(* Logix 5000 project; controller NWGG 1756-L72 rev 35.12; software revision 35.00; part 4 of 19 *)
(* tags used below, declared in another part *)
   DIST_MOVE : ALIAS FOR I3.10;
   DIST_TO_CL : ALIAS FOR I7.2;
   DS_CLEAN_B : ALIAS FOR O13.5;
   DS_DLY_OFF : ALIAS FOR T4[33];
   DS_M : ALIAS FOR O24[1].0;
   DS_M_B : ALIAS FOR B3[101].0;
   DS_MOV_CCW : ALIAS FOR B3[100].13;
   DS_MOV_CW : ALIAS FOR B3[100].12;
   DS_MOVE_SE : ALIAS FOR T4[32];
   DS_POS8 : ALIAS FOR O13.7;
   DS_POS9 : ALIAS FOR O13.8;
   DS_POS_1 : ALIAS FOR I24[0].2;
   DS_POS_10 : ALIAS FOR I24[0].11;
   DS_POS_2 : ALIAS FOR I24[0].3;
   DS_POS_3 : ALIAS FOR I24[0].4;
   DS_POS_4 : ALIAS FOR I24[0].5;
   DS_POS_5 : ALIAS FOR I24[0].6;
   DS_POS_6 : ALIAS FOR I24[0].7;
   DS_POS_7 : ALIAS FOR I24[0].8;
   DS_POS_8 : ALIAS FOR I24[0].9;
   DS_POS_9 : ALIAS FOR I24[0].10;
   DS_SEEK_1 : ALIAS FOR B3[102].1;
   DS_SEEK_10 : ALIAS FOR B3[102].10;
   DS_SEEK_2 : ALIAS FOR B3[102].2;
   DS_SEEK_3 : ALIAS FOR B3[102].3;
   DS_SEEK_4 : ALIAS FOR B3[102].4;
   DS_SEEK_5 : ALIAS FOR B3[102].5;
   DS_SEEK_6 : ALIAS FOR B3[102].6;
   DS_SEEK_7 : ALIAS FOR B3[102].7;
   DS_SEEK_8 : ALIAS FOR B3[102].8;
   DS_SEEK_9 : ALIAS FOR B3[102].9;
   DS_SET_IN : ALIAS FOR N10[0];
   DS_SPOUT_C : ALIAS FOR O24[1].3;
   DS_SPOUT_C1 : ALIAS FOR O24[1].4;
   DS_SPOUT_D : ALIAS FOR I24[0].1;
   DS_SPOUT_D1 : ALIAS FOR O24[1].1;
   DS_SPOUT_D3 : ALIAS FOR B3[101].1;
   DS_SPOUT_U : ALIAS FOR I24[0].0;
   DS_SPOUT_U1 : ALIAS FOR O24[1].2;
   DS_SPOUT_U2 : ALIAS FOR B3[101].2;
   DS_START_M : ALIAS FOR B3[102].11;
   DS_STOP_MO : ALIAS FOR B3[102].0;
   DS_T21 : ALIAS FOR O13.0;
   DS_T22 : ALIAS FOR O13.1;
   DS_T23 : ALIAS FOR O13.9;
   DS_T231 : ALIAS FOR O13.2;
   DS_T24 : ALIAS FOR O13.3;
   DS_T25 : ALIAS FOR O13.4;
   DS_T26 : ALIAS FOR O13.6;
   I24_004_Bit03 : ALIAS FOR I24[4].3;
   I24_004_Bit04 : ALIAS FOR I24[4].4;
   I24_004_Bit05 : ALIAS FOR I24[4].5;
   I24_004_Bit06 : ALIAS FOR I24[4].6;
   I24_004_Bit07 : ALIAS FOR I24[4].7;
   I24_004_Bit08 : ALIAS FOR I24[4].8;
   I24_004_Bit09 : ALIAS FOR I24[4].9;
   I24_004_Bit10 : ALIAS FOR I24[4].10;
   I24_004_Bit11 : ALIAS FOR I24[4].11;
   I24_004_Bit12 : ALIAS FOR I24[4].12;
   I2_000_Bit07 : ALIAS FOR I2.7;
   I2_000_Bit10 : ALIAS FOR I2.10;
   I2_000_Bit13 : ALIAS FOR I2.13;
   I3_000_Bit01 : ALIAS FOR I3.1;
   I3_000_Bit04 : ALIAS FOR I3.4;
   I3_000_Bit07 : ALIAS FOR I3.7;
   O24_005_Bit03 : ALIAS FOR O24[5].3;
   O24_005_Bit04 : ALIAS FOR O24[5].4;
   O24_005_Bit05 : ALIAS FOR O24[5].5;
   O24_005_Bit06 : ALIAS FOR O24[5].6;
   O24_005_Bit07 : ALIAS FOR O24[5].7;
   O24_005_Bit08 : ALIAS FOR O24[5].8;
   O24_005_Bit09 : ALIAS FOR O24[5].9;
   O24_005_Bit10 : ALIAS FOR O24[5].10;
   O24_005_Bit11 : ALIAS FOR O24[5].11;
   O24_005_Bit12 : ALIAS FOR O24[5].12;
   P10_AUTO_S : ALIAS FOR B3[5].10;
   P10_RUN_AU1 : ALIAS FOR B3[4].10;
   P10_SEC_SE : ALIAS FOR B17[1].10;
   P4_RUN_AUT1 : ALIAS FOR B3[4].4;
   P4_SEC_SEL : ALIAS FOR B17[1].4;
   P5_AUTO_SE : ALIAS FOR B3[5].5;
   P5_RUN_AUT1 : ALIAS FOR B3[4].5;
   P5_SEC_SEL : ALIAS FOR B17[1].5;
   P6_AUTO_SE : ALIAS FOR B3[5].6;
   P6_RUN_AUT1 : ALIAS FOR B3[4].6;
   P6_SEC_SEL : ALIAS FOR B17[1].6;
   P7_AUTO_SE : ALIAS FOR B3[5].7;
   P7_RUN_AUT1 : ALIAS FOR B3[4].7;
   P7_SEC_SEL : ALIAS FOR B17[1].7;
   P8_AUTO_SE : ALIAS FOR B3[5].8;
   P8_RUN_AUT1 : ALIAS FOR B3[4].8;
   P8_SEC_SEL : ALIAS FOR B17[1].8;
   P_RESET_AU : ALIAS FOR B3[4].0;
   SYMBOL_ANA : ALIAS FOR N10[1];
   T11_TREAT : ALIAS FOR B3[11].0;
   T12_TREAT : ALIAS FOR B3[12].0;
   T13_TREAT : ALIAS FOR B3[13].0;
   T13C_TREAT : ALIAS FOR B21[70].10;
   T14_TREAT : ALIAS FOR B3[14].0;
   T15_TREAT : ALIAS FOR B3[15].0;
   T16_TREAT : ALIAS FOR B3[16].0;
   T17_TREAT : ALIAS FOR B3[17].0;
   T19C_TREAT : ALIAS FOR B21[71].10;
   T21_TREAT : ALIAS FOR B3[21].0;
   T22_TREAT : ALIAS FOR B3[22].0;
   T23_TREAT : ALIAS FOR B3[23].0;
   T24_TREAT : ALIAS FOR B3[24].0;
   T25_TREAT : ALIAS FOR B3[25].0;
   T26_TREAT : ALIAS FOR B3[26].0;
   T27_TREAT : ALIAS FOR B3[27].0;
   T28_TREAT : ALIAS FOR B3[28].0;
   T29_TREAT : ALIAS FOR B3[29].0;
(* _2_MAIN, continued *)

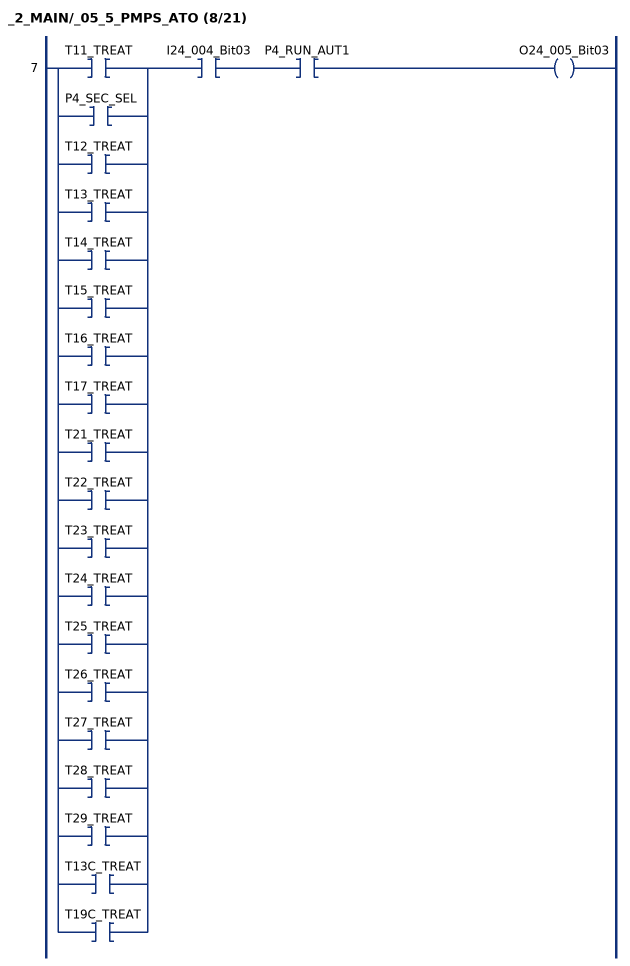
   [picture p56: _2_MAIN/_05_5_PMPS_ATO rungs 7-7]
   7: [XIC(T11_TREAT) ,XIC(P4_SEC_SEL) ,XIC(T12_TREAT) ,XIC(T13_TREAT) ,XIC(T14_TREAT) ,XIC(T15_TREAT) ,XIC(T16_TREAT) ,XIC(T17_TREAT) ,XIC(T21_TREAT) ,XIC(T22_TREAT) ,XIC(T23_TREAT) ,XIC(T24_TREAT) ,XIC(T25_TREAT) ,XIC(T26_TREAT) ,XIC(T27_TREAT) ,XIC(T28_TREAT) ,XIC(T29_TREAT) ,XIC(T13C_TREAT) ,XIC(T19C_TREAT) ]XIC(I24_004_Bit03)XIC(P4_RUN_AUT1)OTE(O24_005_Bit03);
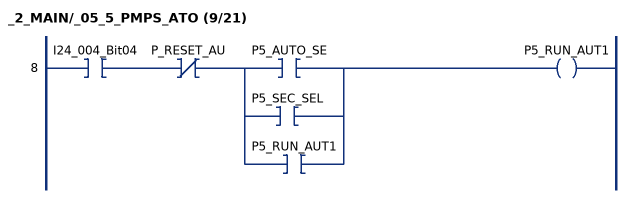
   8: XIC(I24_004_Bit04)XIO(P_RESET_AU)[XIC(P5_AUTO_SE) ,XIC(P5_SEC_SEL) ,XIC(P5_RUN_AUT1) ]OTE(P5_RUN_AUT1);
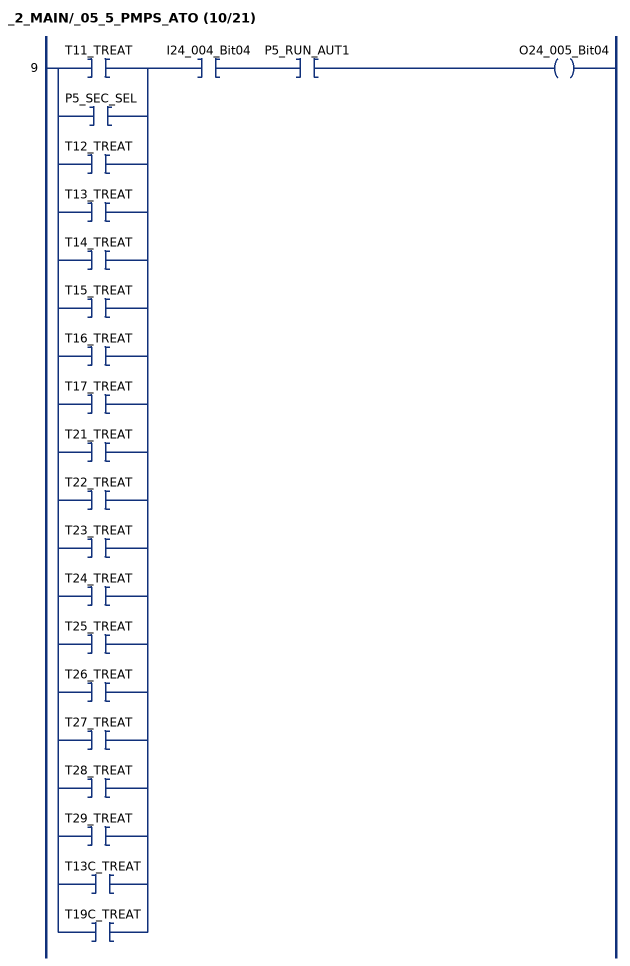
   9: [XIC(T11_TREAT) ,XIC(P5_SEC_SEL) ,XIC(T12_TREAT) ,XIC(T13_TREAT) ,XIC(T14_TREAT) ,XIC(T15_TREAT) ,XIC(T16_TREAT) ,XIC(T17_TREAT) ,XIC(T21_TREAT) ,XIC(T22_TREAT) ,XIC(T23_TREAT) ,XIC(T24_TREAT) ,XIC(T25_TREAT) ,XIC(T26_TREAT) ,XIC(T27_TREAT) ,XIC(T28_TREAT) ,XIC(T29_TREAT) ,XIC(T13C_TREAT) ,XIC(T19C_TREAT) ]XIC(I24_004_Bit04)XIC(P5_RUN_AUT1)OTE(O24_005_Bit04);
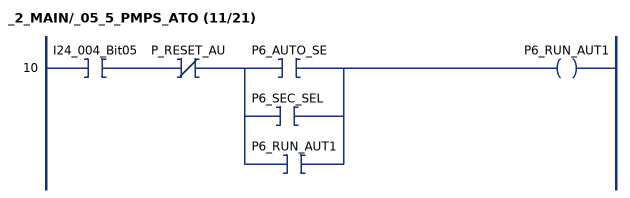
   10: XIC(I24_004_Bit05)XIO(P_RESET_AU)[XIC(P6_AUTO_SE) ,XIC(P6_SEC_SEL) ,XIC(P6_RUN_AUT1) ]OTE(P6_RUN_AUT1);
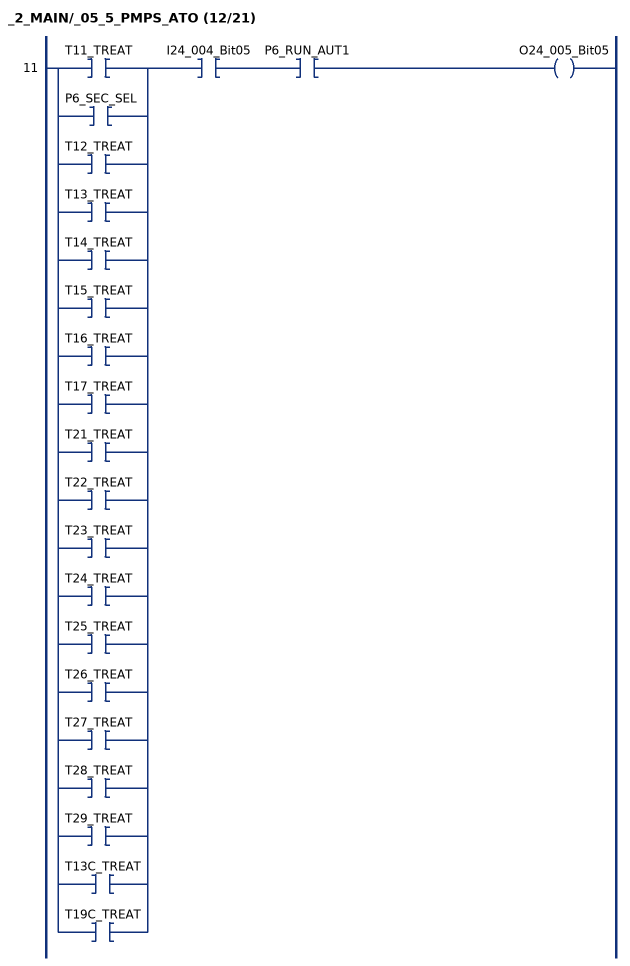
   11: [XIC(T11_TREAT) ,XIC(P6_SEC_SEL) ,XIC(T12_TREAT) ,XIC(T13_TREAT) ,XIC(T14_TREAT) ,XIC(T15_TREAT) ,XIC(T16_TREAT) ,XIC(T17_TREAT) ,XIC(T21_TREAT) ,XIC(T22_TREAT) ,XIC(T23_TREAT) ,XIC(T24_TREAT) ,XIC(T25_TREAT) ,XIC(T26_TREAT) ,XIC(T27_TREAT) ,XIC(T28_TREAT) ,XIC(T29_TREAT) ,XIC(T13C_TREAT) ,XIC(T19C_TREAT) ]XIC(I24_004_Bit05)XIC(P6_RUN_AUT1)OTE(O24_005_Bit05);
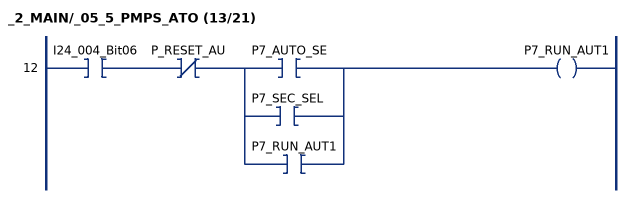
   12: XIC(I24_004_Bit06)XIO(P_RESET_AU)[XIC(P7_AUTO_SE) ,XIC(P7_SEC_SEL) ,XIC(P7_RUN_AUT1) ]OTE(P7_RUN_AUT1);
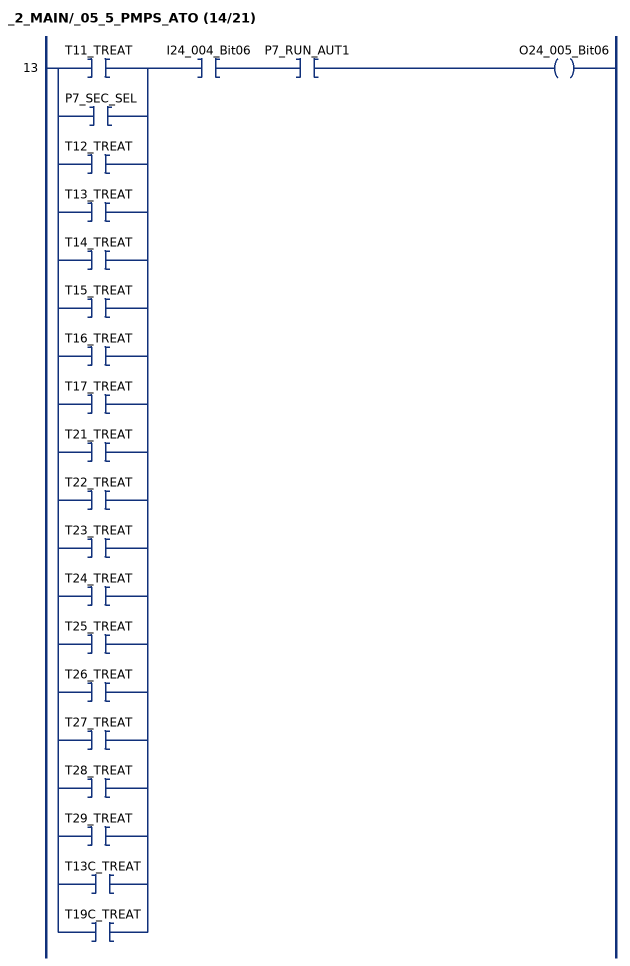
   13: [XIC(T11_TREAT) ,XIC(P7_SEC_SEL) ,XIC(T12_TREAT) ,XIC(T13_TREAT) ,XIC(T14_TREAT) ,XIC(T15_TREAT) ,XIC(T16_TREAT) ,XIC(T17_TREAT) ,XIC(T21_TREAT) ,XIC(T22_TREAT) ,XIC(T23_TREAT) ,XIC(T24_TREAT) ,XIC(T25_TREAT) ,XIC(T26_TREAT) ,XIC(T27_TREAT) ,XIC(T28_TREAT) ,XIC(T29_TREAT) ,XIC(T13C_TREAT) ,XIC(T19C_TREAT) ]XIC(I24_004_Bit06)XIC(P7_RUN_AUT1)OTE(O24_005_Bit06);
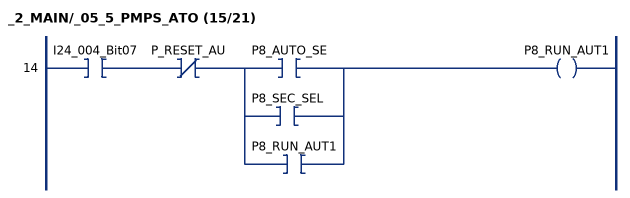
   14: XIC(I24_004_Bit07)XIO(P_RESET_AU)[XIC(P8_AUTO_SE) ,XIC(P8_SEC_SEL) ,XIC(P8_RUN_AUT1) ]OTE(P8_RUN_AUT1);
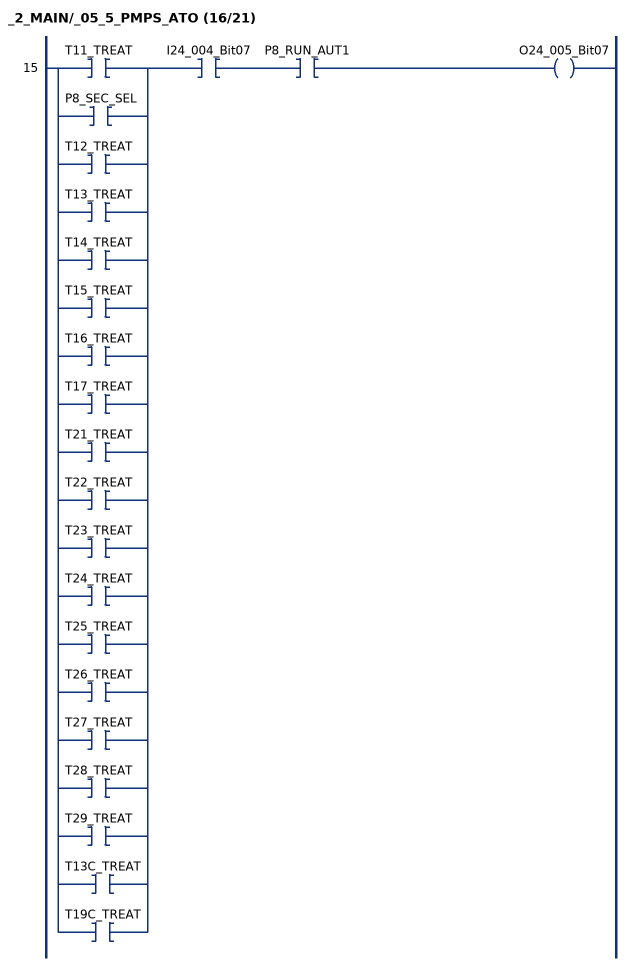
   15: [XIC(T11_TREAT) ,XIC(P8_SEC_SEL) ,XIC(T12_TREAT) ,XIC(T13_TREAT) ,XIC(T14_TREAT) ,XIC(T15_TREAT) ,XIC(T16_TREAT) ,XIC(T17_TREAT) ,XIC(T21_TREAT) ,XIC(T22_TREAT) ,XIC(T23_TREAT) ,XIC(T24_TREAT) ,XIC(T25_TREAT) ,XIC(T26_TREAT) ,XIC(T27_TREAT) ,XIC(T28_TREAT) ,XIC(T29_TREAT) ,XIC(T13C_TREAT) ,XIC(T19C_TREAT) ]XIC(I24_004_Bit07)XIC(P8_RUN_AUT1)OTE(O24_005_Bit07);
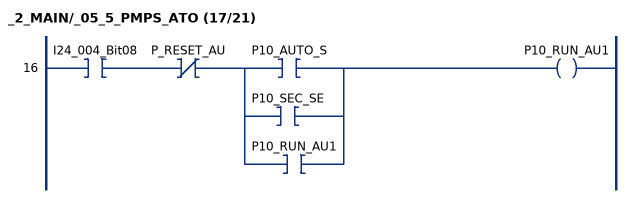
   16: XIC(I24_004_Bit08)XIO(P_RESET_AU)[XIC(P10_AUTO_S) ,XIC(P10_SEC_SE) ,XIC(P10_RUN_AU1) ]OTE(P10_RUN_AU1);
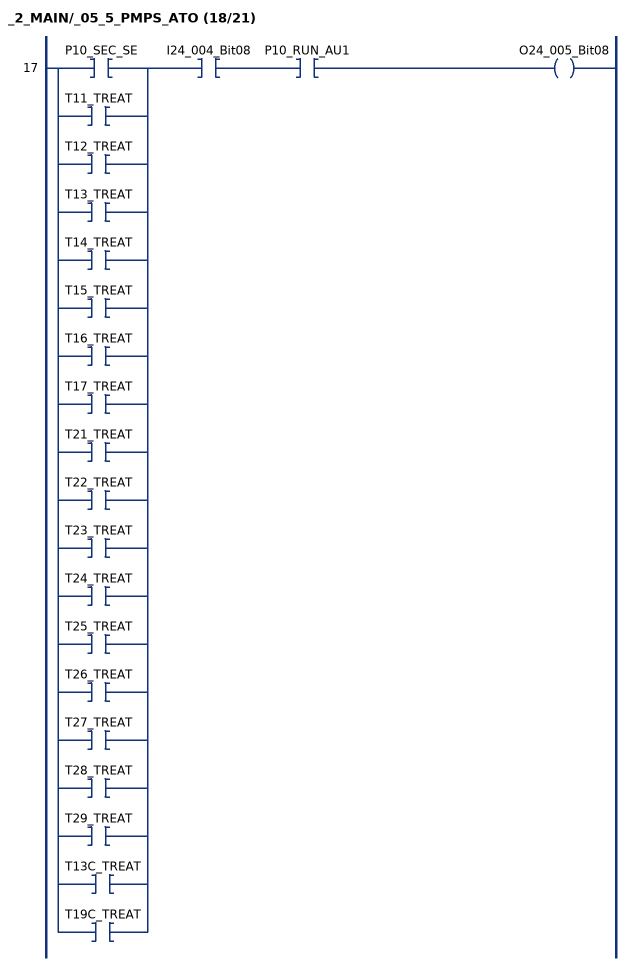
   17: [XIC(P10_SEC_SE) ,XIC(T11_TREAT) ,XIC(T12_TREAT) ,XIC(T13_TREAT) ,XIC(T14_TREAT) ,XIC(T15_TREAT) ,XIC(T16_TREAT) ,XIC(T17_TREAT) ,XIC(T21_TREAT) ,XIC(T22_TREAT) ,XIC(T23_TREAT) ,XIC(T24_TREAT) ,XIC(T25_TREAT) ,XIC(T26_TREAT) ,XIC(T27_TREAT) ,XIC(T28_TREAT) ,XIC(T29_TREAT) ,XIC(T13C_TREAT) ,XIC(T19C_TREAT) ]XIC(I24_004_Bit08)XIC(P10_RUN_AU1)OTE(O24_005_Bit08);
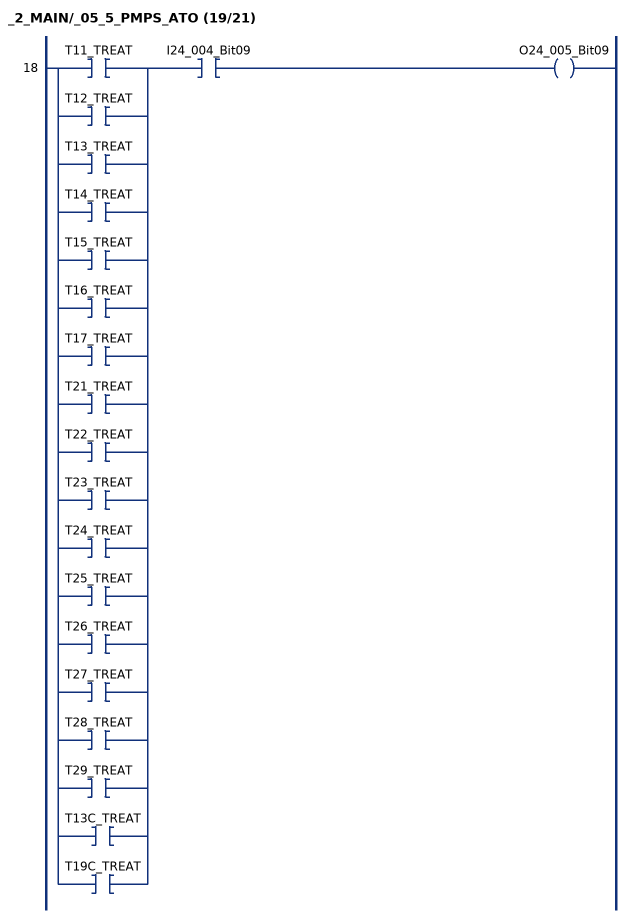
   18: [XIC(T11_TREAT) ,XIC(T12_TREAT) ,XIC(T13_TREAT) ,XIC(T14_TREAT) ,XIC(T15_TREAT) ,XIC(T16_TREAT) ,XIC(T17_TREAT) ,XIC(T21_TREAT) ,XIC(T22_TREAT) ,XIC(T23_TREAT) ,XIC(T24_TREAT) ,XIC(T25_TREAT) ,XIC(T26_TREAT) ,XIC(T27_TREAT) ,XIC(T28_TREAT) ,XIC(T29_TREAT) ,XIC(T13C_TREAT) ,XIC(T19C_TREAT) ]XIC(I24_004_Bit09)OTE(O24_005_Bit09);
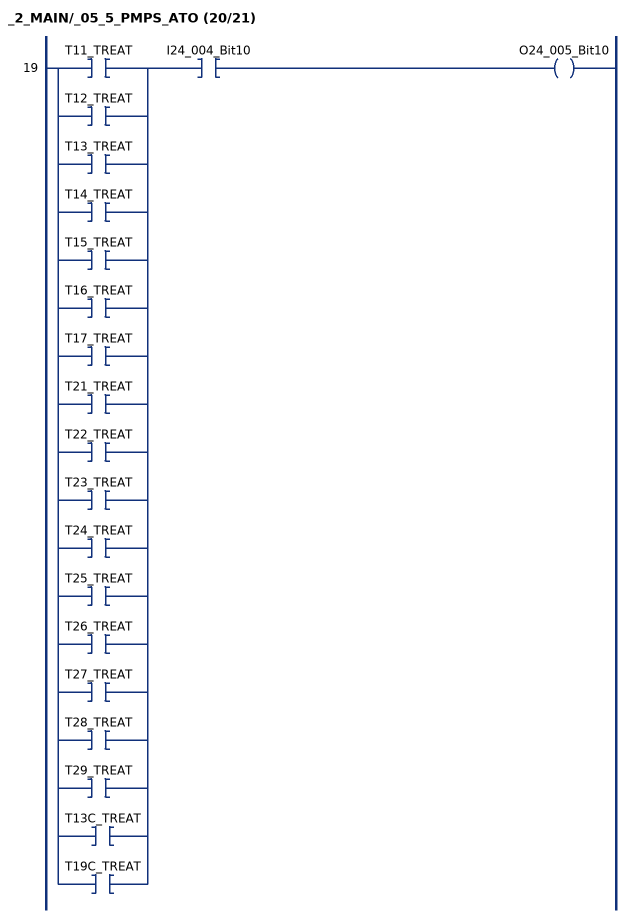
   19: [XIC(T11_TREAT) ,XIC(T12_TREAT) ,XIC(T13_TREAT) ,XIC(T14_TREAT) ,XIC(T15_TREAT) ,XIC(T16_TREAT) ,XIC(T17_TREAT) ,XIC(T21_TREAT) ,XIC(T22_TREAT) ,XIC(T23_TREAT) ,XIC(T24_TREAT) ,XIC(T25_TREAT) ,XIC(T26_TREAT) ,XIC(T27_TREAT) ,XIC(T28_TREAT) ,XIC(T29_TREAT) ,XIC(T13C_TREAT) ,XIC(T19C_TREAT) ]XIC(I24_004_Bit10)OTE(O24_005_Bit10);
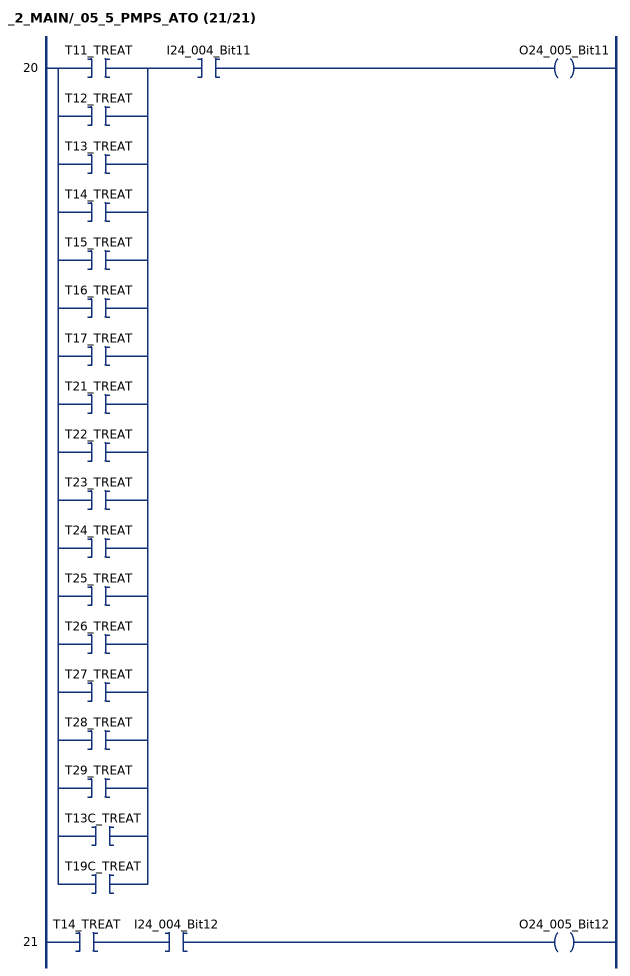
   20: [XIC(T11_TREAT) ,XIC(T12_TREAT) ,XIC(T13_TREAT) ,XIC(T14_TREAT) ,XIC(T15_TREAT) ,XIC(T16_TREAT) ,XIC(T17_TREAT) ,XIC(T21_TREAT) ,XIC(T22_TREAT) ,XIC(T23_TREAT) ,XIC(T24_TREAT) ,XIC(T25_TREAT) ,XIC(T26_TREAT) ,XIC(T27_TREAT) ,XIC(T28_TREAT) ,XIC(T29_TREAT) ,XIC(T13C_TREAT) ,XIC(T19C_TREAT) ]XIC(I24_004_Bit11)OTE(O24_005_Bit11);
   21: XIC(T14_TREAT)XIC(I24_004_Bit12)OTE(O24_005_Bit12);
END_ROUTINE

ROUTINE _06_DISTRIB_SW   (* ladder *)
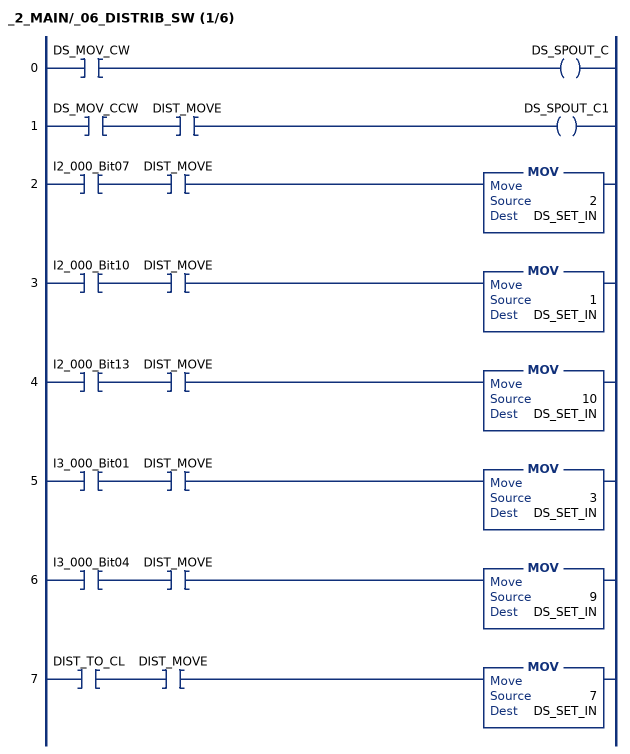
   0: XIC(DS_MOV_CW)OTE(DS_SPOUT_C);
   1: XIC(DS_MOV_CCW)XIC(DIST_MOVE)OTE(DS_SPOUT_C1);
   2: XIC(I2_000_Bit07)XIC(DIST_MOVE)MOV(2,DS_SET_IN);
   3: XIC(I2_000_Bit10)XIC(DIST_MOVE)MOV(1,DS_SET_IN);
   4: XIC(I2_000_Bit13)XIC(DIST_MOVE)MOV(10,DS_SET_IN);
   5: XIC(I3_000_Bit01)XIC(DIST_MOVE)MOV(3,DS_SET_IN);
   6: XIC(I3_000_Bit04)XIC(DIST_MOVE)MOV(9,DS_SET_IN);
   7: XIC(DIST_TO_CL)XIC(DIST_MOVE)MOV(7,DS_SET_IN);
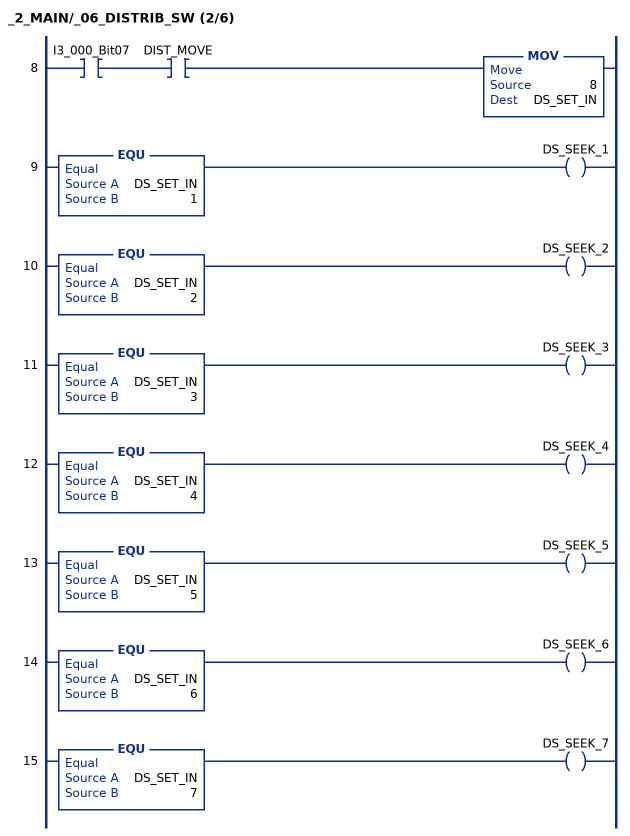
   8: XIC(I3_000_Bit07)XIC(DIST_MOVE)MOV(8,DS_SET_IN);
   9: EQU(DS_SET_IN,1)OTE(DS_SEEK_1);
   10: EQU(DS_SET_IN,2)OTE(DS_SEEK_2);
   11: EQU(DS_SET_IN,3)OTE(DS_SEEK_3);
   12: EQU(DS_SET_IN,4)OTE(DS_SEEK_4);
   13: EQU(DS_SET_IN,5)OTE(DS_SEEK_5);
   14: EQU(DS_SET_IN,6)OTE(DS_SEEK_6);
   15: EQU(DS_SET_IN,7)OTE(DS_SEEK_7);
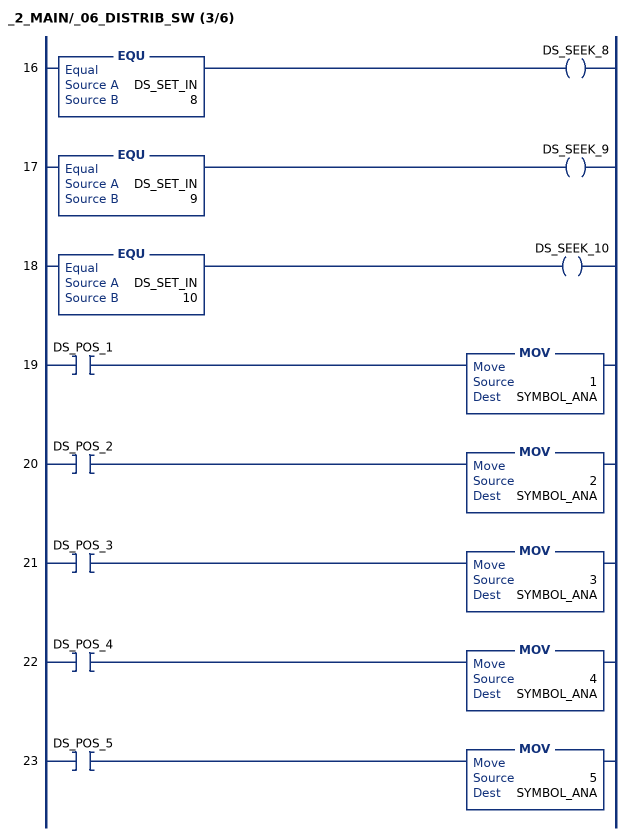
   16: EQU(DS_SET_IN,8)OTE(DS_SEEK_8);
   17: EQU(DS_SET_IN,9)OTE(DS_SEEK_9);
   18: EQU(DS_SET_IN,10)OTE(DS_SEEK_10);
   19: XIC(DS_POS_1)MOV(1,SYMBOL_ANA);
   20: XIC(DS_POS_2)MOV(2,SYMBOL_ANA);
   21: XIC(DS_POS_3)MOV(3,SYMBOL_ANA);
   22: XIC(DS_POS_4)MOV(4,SYMBOL_ANA);
   23: XIC(DS_POS_5)MOV(5,SYMBOL_ANA);
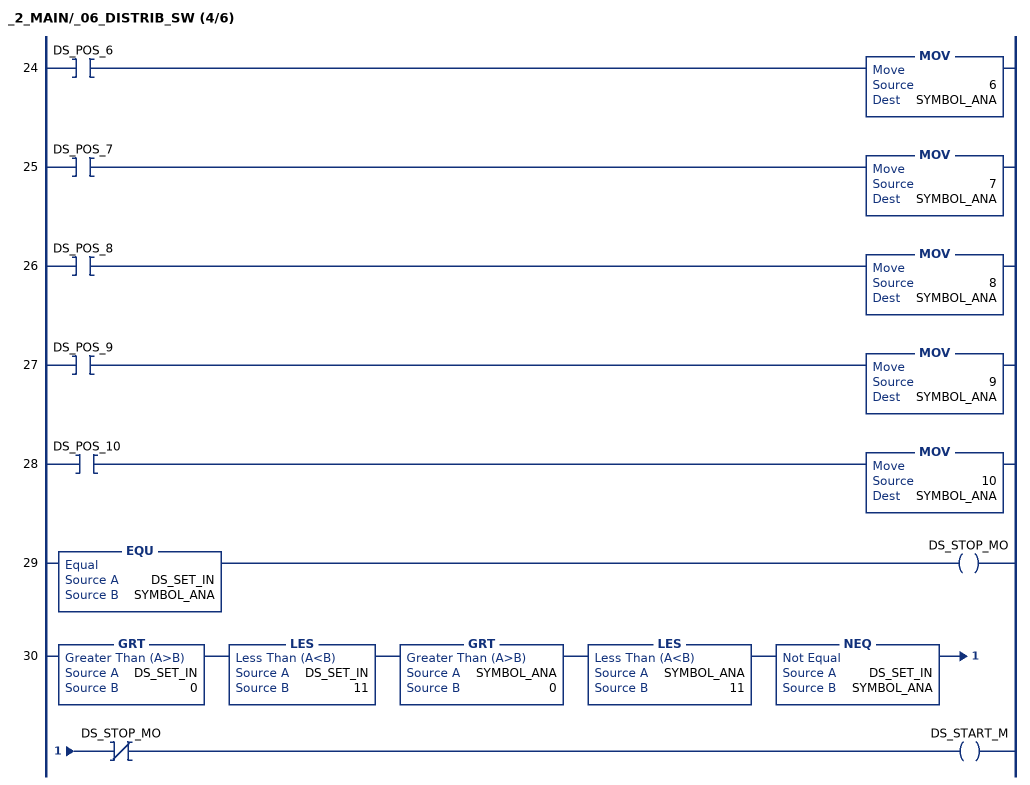
   24: XIC(DS_POS_6)MOV(6,SYMBOL_ANA);
   25: XIC(DS_POS_7)MOV(7,SYMBOL_ANA);
   26: XIC(DS_POS_8)MOV(8,SYMBOL_ANA);
   27: XIC(DS_POS_9)MOV(9,SYMBOL_ANA);
   28: XIC(DS_POS_10)MOV(10,SYMBOL_ANA);
   29: EQU(DS_SET_IN,SYMBOL_ANA)OTE(DS_STOP_MO);
   30: GRT(DS_SET_IN,0)LES(DS_SET_IN,11)GRT(SYMBOL_ANA,0)LES(SYMBOL_ANA,11)NEQ(DS_SET_IN,SYMBOL_ANA)XIO(DS_STOP_MO)OTE(DS_START_M);
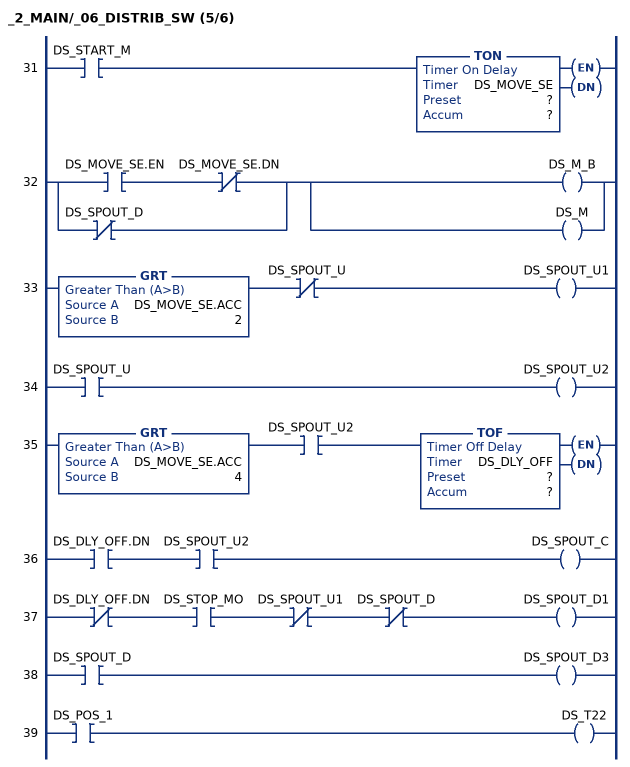
   31: XIC(DS_START_M)TON(DS_MOVE_SE,?,?);
   32: [XIC(DS_MOVE_SE.EN) XIO(DS_MOVE_SE.DN) ,XIO(DS_SPOUT_D) ][OTE(DS_M_B) ,OTE(DS_M) ];
   33: GRT(DS_MOVE_SE.ACC,2)XIO(DS_SPOUT_U)OTE(DS_SPOUT_U1);
   34: XIC(DS_SPOUT_U)OTE(DS_SPOUT_U2);
   35: GRT(DS_MOVE_SE.ACC,4)XIC(DS_SPOUT_U2)TOF(DS_DLY_OFF,?,?);
   36: XIC(DS_DLY_OFF.DN)XIC(DS_SPOUT_U2)OTE(DS_SPOUT_C);
   37: XIO(DS_DLY_OFF.DN)XIC(DS_STOP_MO)XIO(DS_SPOUT_U1)XIO(DS_SPOUT_D)OTE(DS_SPOUT_D1);
   38: XIC(DS_SPOUT_D)OTE(DS_SPOUT_D3);
   39: XIC(DS_POS_1)OTE(DS_T22);
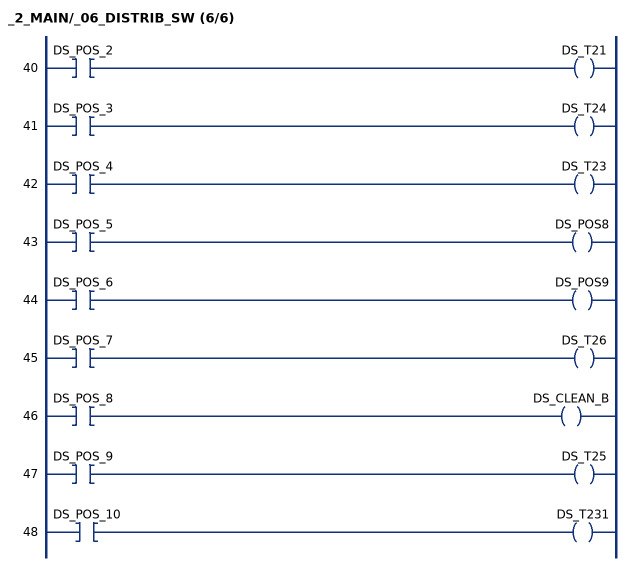
   40: XIC(DS_POS_2)OTE(DS_T21);
   41: XIC(DS_POS_3)OTE(DS_T24);
   42: XIC(DS_POS_4)OTE(DS_T23);
   43: XIC(DS_POS_5)OTE(DS_POS8);
   44: XIC(DS_POS_6)OTE(DS_POS9);
   45: XIC(DS_POS_7)OTE(DS_T26);
   46: XIC(DS_POS_8)OTE(DS_CLEAN_B);
   47: XIC(DS_POS_9)OTE(DS_T25);
   48: XIC(DS_POS_10)OTE(DS_T231);
END_ROUTINE
